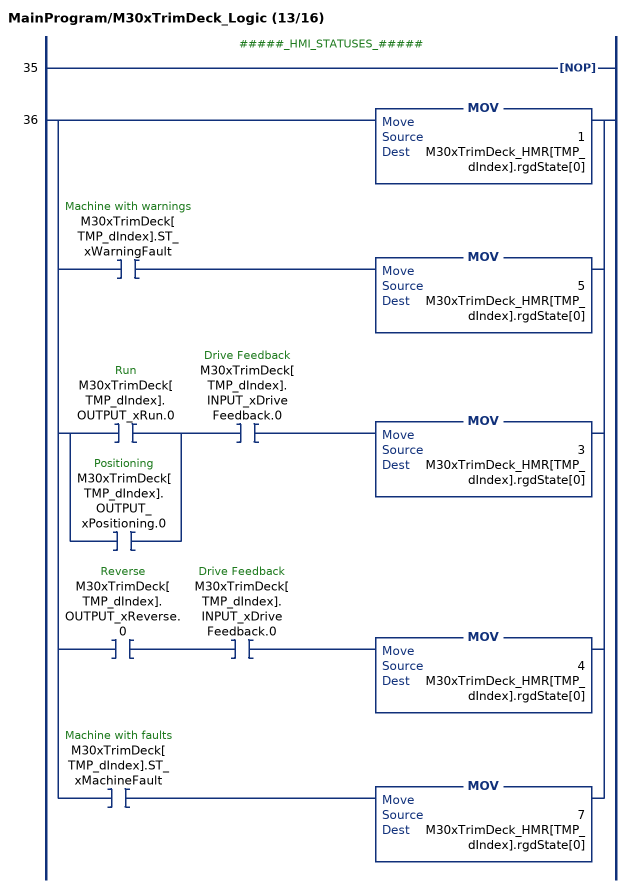
   // #####_HMI_STATUSES_#####
   35: NOP();
   36: [MOV(1,M30xTrimDeck_HMR[TMP_dIndex].rgdState[0]) ,XIC(M30xTrimDeck[TMP_dIndex].ST_xWarningFault) MOV(5,M30xTrimDeck_HMR[TMP_dIndex].rgdState[0]) ,[XIC(M30xTrimDeck[TMP_dIndex].OUTPUT_xRun.0) ,XIC(M30xTrimDeck[TMP_dIndex].OUTPUT_xPositioning.0) ] XIC(M30xTrimDeck[TMP_dIndex].INPUT_xDriveFeedback.0) MOV(3,M30xTrimDeck_HMR[TMP_dIndex].rgdState[0]) ,XIC(M30xTrimDeck[TMP_dIndex].OUTPUT_xReverse.0) XIC(M30xTrimDeck[TMP_dIndex].INPUT_xDriveFeedback.0) MOV(4,M30xTrimDeck_HMR[TMP_dIndex].rgdState[0]) ,XIC(M30xTrimDeck[TMP_dIndex].ST_xMachineFault) MOV(7,M30xTrimDeck_HMR[TMP_dIndex].rgdState[0]) ];
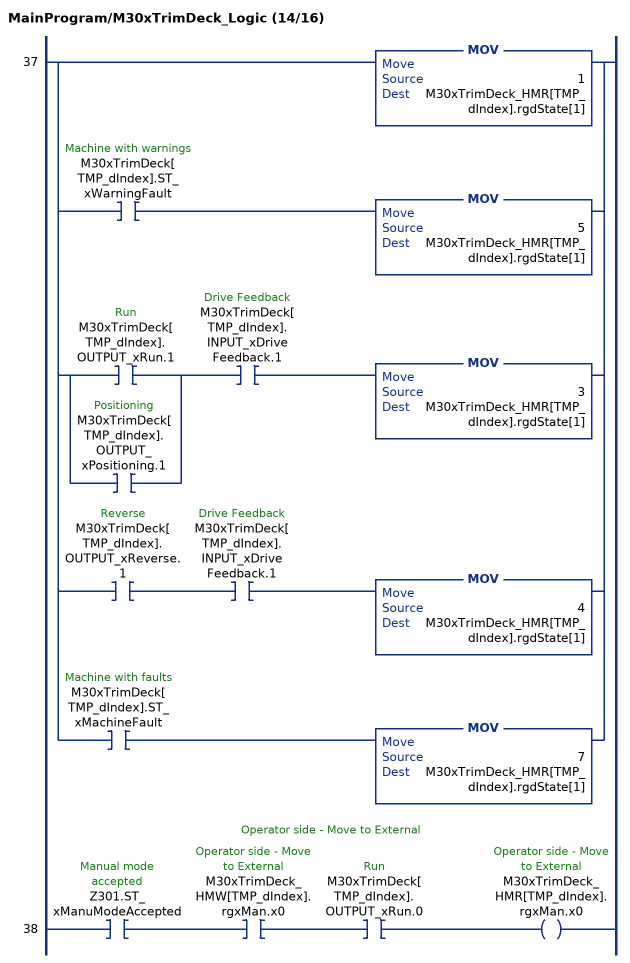
   37: [MOV(1,M30xTrimDeck_HMR[TMP_dIndex].rgdState[1]) ,XIC(M30xTrimDeck[TMP_dIndex].ST_xWarningFault) MOV(5,M30xTrimDeck_HMR[TMP_dIndex].rgdState[1]) ,[XIC(M30xTrimDeck[TMP_dIndex].OUTPUT_xRun.1) ,XIC(M30xTrimDeck[TMP_dIndex].OUTPUT_xPositioning.1) ] XIC(M30xTrimDeck[TMP_dIndex].INPUT_xDriveFeedback.1) MOV(3,M30xTrimDeck_HMR[TMP_dIndex].rgdState[1]) ,XIC(M30xTrimDeck[TMP_dIndex].OUTPUT_xReverse.1) XIC(M30xTrimDeck[TMP_dIndex].INPUT_xDriveFeedback.1) MOV(4,M30xTrimDeck_HMR[TMP_dIndex].rgdState[1]) ,XIC(M30xTrimDeck[TMP_dIndex].ST_xMachineFault) MOV(7,M30xTrimDeck_HMR[TMP_dIndex].rgdState[1]) ];
   // Operator side - Move to External
   38: XIC(Z301.ST_xManuModeAccepted)XIC(M30xTrimDeck_HMW[TMP_dIndex].rgxMan.x0)XIC(M30xTrimDeck[TMP_dIndex].OUTPUT_xRun.0)OTE(M30xTrimDeck_HMR[TMP_dIndex].rgxMan.x0);
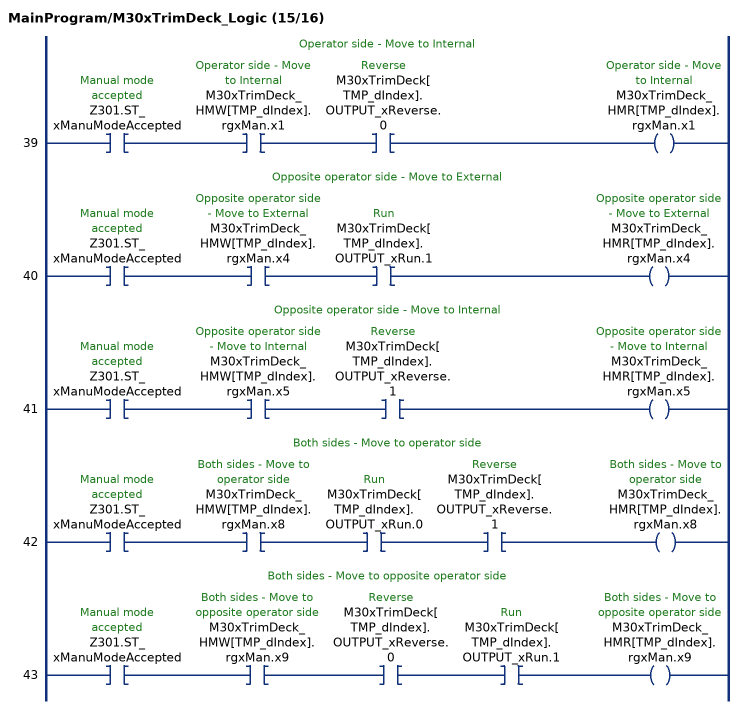
   // Operator side - Move to Internal
   39: XIC(Z301.ST_xManuModeAccepted)XIC(M30xTrimDeck_HMW[TMP_dIndex].rgxMan.x1)XIC(M30xTrimDeck[TMP_dIndex].OUTPUT_xReverse.0)OTE(M30xTrimDeck_HMR[TMP_dIndex].rgxMan.x1);
   // Opposite operator side - Move to External
   40: XIC(Z301.ST_xManuModeAccepted)XIC(M30xTrimDeck_HMW[TMP_dIndex].rgxMan.x4)XIC(M30xTrimDeck[TMP_dIndex].OUTPUT_xRun.1)OTE(M30xTrimDeck_HMR[TMP_dIndex].rgxMan.x4);
   // Opposite operator side - Move to Internal
   41: XIC(Z301.ST_xManuModeAccepted)XIC(M30xTrimDeck_HMW[TMP_dIndex].rgxMan.x5)XIC(M30xTrimDeck[TMP_dIndex].OUTPUT_xReverse.1)OTE(M30xTrimDeck_HMR[TMP_dIndex].rgxMan.x5);
   // Both sides - Move to operator side
   42: XIC(Z301.ST_xManuModeAccepted)XIC(M30xTrimDeck_HMW[TMP_dIndex].rgxMan.x8)XIC(M30xTrimDeck[TMP_dIndex].OUTPUT_xRun.0)XIC(M30xTrimDeck[TMP_dIndex].OUTPUT_xReverse.1)OTE(M30xTrimDeck_HMR[TMP_dIndex].rgxMan.x8);
   // Both sides - Move to opposite operator side
   43: XIC(Z301.ST_xManuModeAccepted)XIC(M30xTrimDeck_HMW[TMP_dIndex].rgxMan.x9)XIC(M30xTrimDeck[TMP_dIndex].OUTPUT_xReverse.0)XIC(M30xTrimDeck[TMP_dIndex].OUTPUT_xRun.1)OTE(M30xTrimDeck_HMR[TMP_dIndex].rgxMan.x9);
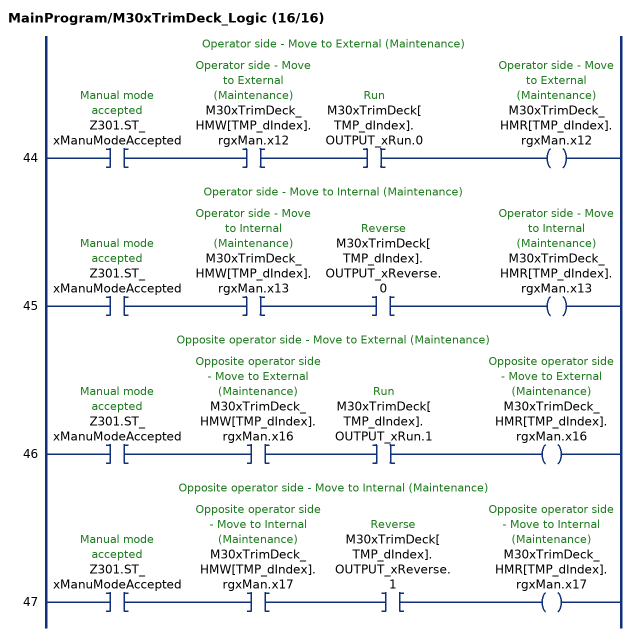
   // Operator side - Move to External (Maintenance)
   44: XIC(Z301.ST_xManuModeAccepted)XIC(M30xTrimDeck_HMW[TMP_dIndex].rgxMan.x12)XIC(M30xTrimDeck[TMP_dIndex].OUTPUT_xRun.0)OTE(M30xTrimDeck_HMR[TMP_dIndex].rgxMan.x12);
   // Operator side - Move to Internal (Maintenance)
   45: XIC(Z301.ST_xManuModeAccepted)XIC(M30xTrimDeck_HMW[TMP_dIndex].rgxMan.x13)XIC(M30xTrimDeck[TMP_dIndex].OUTPUT_xReverse.0)OTE(M30xTrimDeck_HMR[TMP_dIndex].rgxMan.x13);
   // Opposite operator side - Move to External (Maintenance)
   46: XIC(Z301.ST_xManuModeAccepted)XIC(M30xTrimDeck_HMW[TMP_dIndex].rgxMan.x16)XIC(M30xTrimDeck[TMP_dIndex].OUTPUT_xRun.1)OTE(M30xTrimDeck_HMR[TMP_dIndex].rgxMan.x16);
   // Opposite operator side - Move to Internal (Maintenance)
   47: XIC(Z301.ST_xManuModeAccepted)XIC(M30xTrimDeck_HMW[TMP_dIndex].rgxMan.x17)XIC(M30xTrimDeck[TMP_dIndex].OUTPUT_xReverse.1)OTE(M30xTrimDeck_HMR[TMP_dIndex].rgxMan.x17);
END_ROUTINE

ROUTINE M30xTrimDeckManagement   (* ladder *)
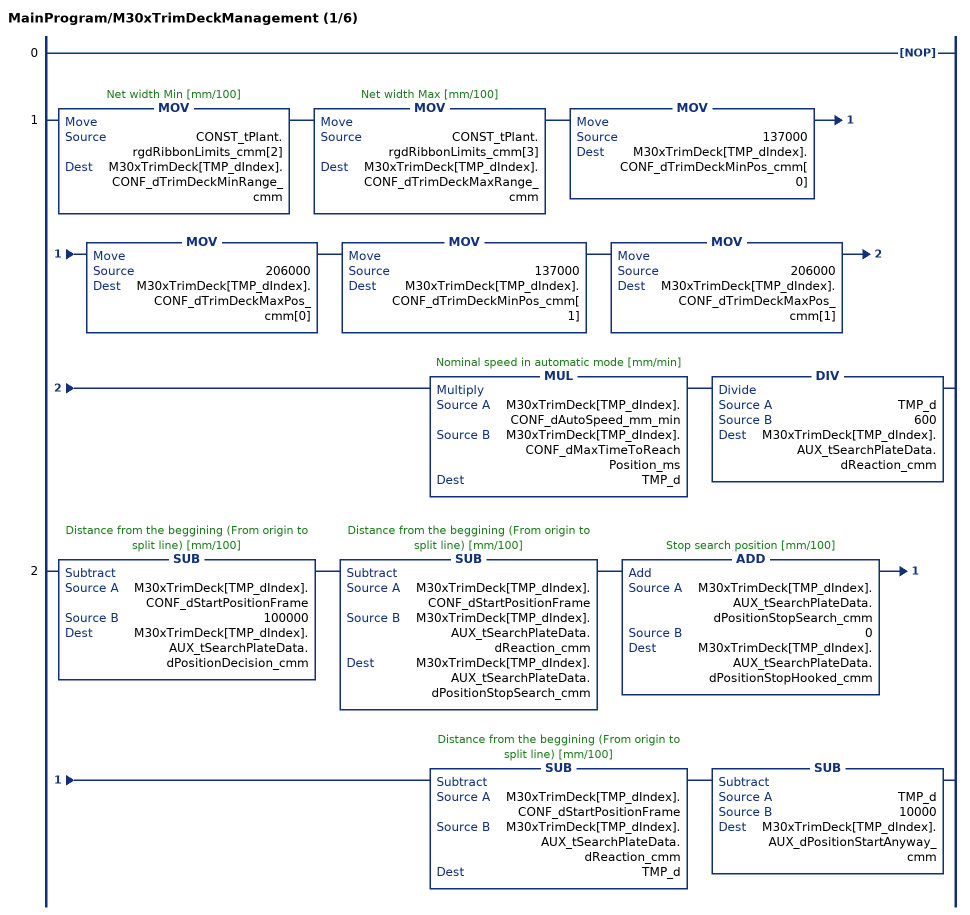
   0: NOP();
   1: MOV(CONST_tPlant.rgdRibbonLimits_cmm[2],M30xTrimDeck[TMP_dIndex].CONF_dTrimDeckMinRange_cmm)MOV(CONST_tPlant.rgdRibbonLimits_cmm[3],M30xTrimDeck[TMP_dIndex].CONF_dTrimDeckMaxRange_cmm)MOV(137000,M30xTrimDeck[TMP_dIndex].CONF_dTrimDeckMinPos_cmm[0])MOV(206000,M30xTrimDeck[TMP_dIndex].CONF_dTrimDeckMaxPos_cmm[0])MOV(137000,M30xTrimDeck[TMP_dIndex].CONF_dTrimDeckMinPos_cmm[1])MOV(206000,M30xTrimDeck[TMP_dIndex].CONF_dTrimDeckMaxPos_cmm[1])MUL(M30xTrimDeck[TMP_dIndex].CONF_dAutoSpeed_mm_min,M30xTrimDeck[TMP_dIndex].CONF_dMaxTimeToReachPosition_ms,TMP_d)DIV(TMP_d,600,M30xTrimDeck[TMP_dIndex].AUX_tSearchPlateData.dReaction_cmm);
   2: SUB(M30xTrimDeck[TMP_dIndex].CONF_dStartPositionFrame,100000,M30xTrimDeck[TMP_dIndex].AUX_tSearchPlateData.dPositionDecision_cmm)SUB(M30xTrimDeck[TMP_dIndex].CONF_dStartPositionFrame,M30xTrimDeck[TMP_dIndex].AUX_tSearchPlateData.dReaction_cmm,M30xTrimDeck[TMP_dIndex].AUX_tSearchPlateData.dPositionStopSearch_cmm)ADD(M30xTrimDeck[TMP_dIndex].AUX_tSearchPlateData.dPositionStopSearch_cmm,0,M30xTrimDeck[TMP_dIndex].AUX_tSearchPlateData.dPositionStopHooked_cmm)SUB(M30xTrimDeck[TMP_dIndex].CONF_dStartPositionFrame,M30xTrimDeck[TMP_dIndex].AUX_tSearchPlateData.dReaction_cmm,TMP_d)SUB(TMP_d,10000,M30xTrimDeck[TMP_dIndex].AUX_dPositionStartAnyway_cmm);
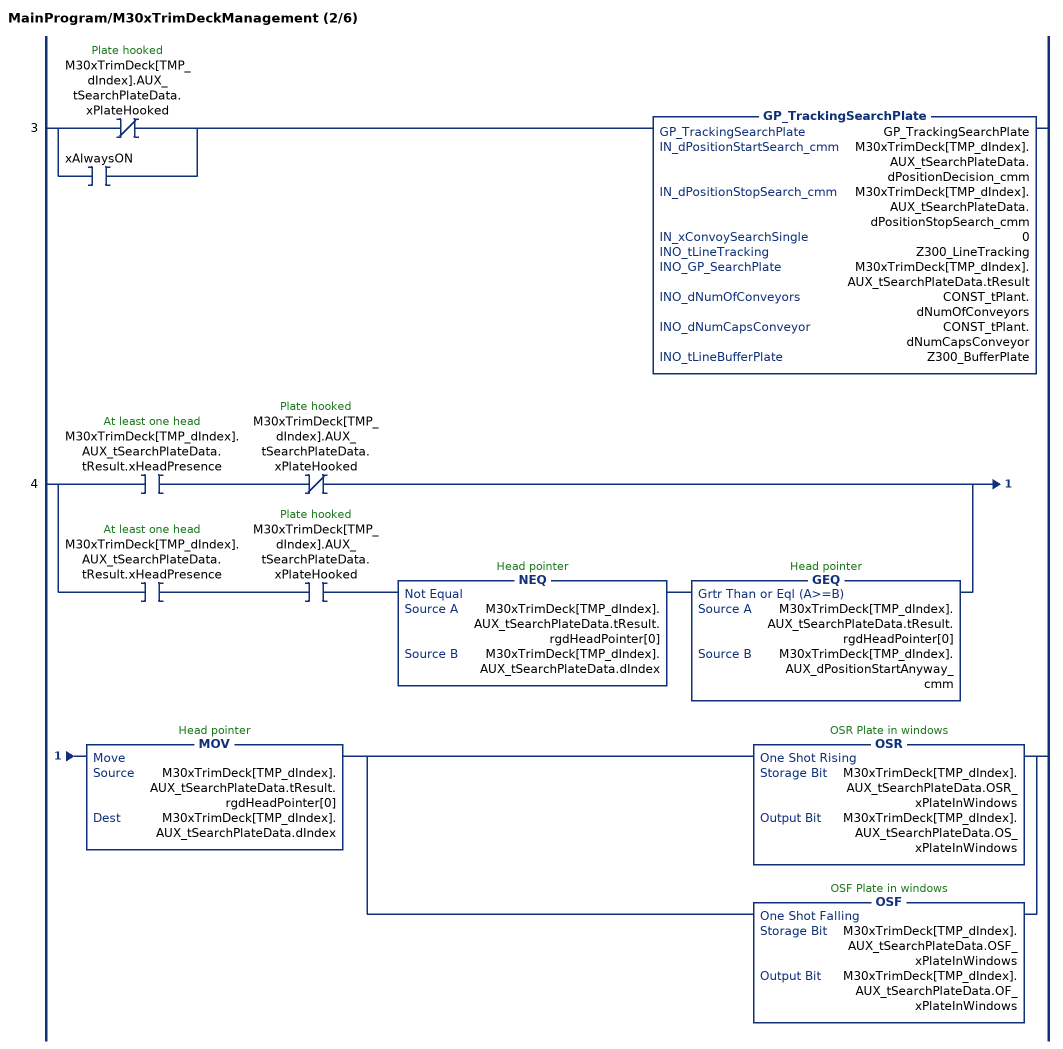
   3: [XIO(M30xTrimDeck[TMP_dIndex].AUX_tSearchPlateData.xPlateHooked) ,XIC(xAlwaysON) ]GP_TrackingSearchPlate(GP_TrackingSearchPlate,M30xTrimDeck[TMP_dIndex].AUX_tSearchPlateData.dPositionDecision_cmm,M30xTrimDeck[TMP_dIndex].AUX_tSearchPlateData.dPositionStopSearch_cmm,0,Z300_LineTracking,M30xTrimDeck[TMP_dIndex].AUX_tSearchPlateData.tResult,CONST_tPlant.dNumOfConveyors,CONST_tPlant.dNumCapsConveyor,Z300_BufferPlate);
   4: [XIC(M30xTrimDeck[TMP_dIndex].AUX_tSearchPlateData.tResult.xHeadPresence) XIO(M30xTrimDeck[TMP_dIndex].AUX_tSearchPlateData.xPlateHooked) ,XIC(M30xTrimDeck[TMP_dIndex].AUX_tSearchPlateData.tResult.xHeadPresence) XIC(M30xTrimDeck[TMP_dIndex].AUX_tSearchPlateData.xPlateHooked) NEQ(M30xTrimDeck[TMP_dIndex].AUX_tSearchPlateData.tResult.rgdHeadPointer[0],M30xTrimDeck[TMP_dIndex].AUX_tSearchPlateData.dIndex) GEQ(M30xTrimDeck[TMP_dIndex].AUX_tSearchPlateData.tResult.rgdHeadPointer[0],M30xTrimDeck[TMP_dIndex].AUX_dPositionStartAnyway_cmm) ]MOV(M30xTrimDeck[TMP_dIndex].AUX_tSearchPlateData.tResult.rgdHeadPointer[0],M30xTrimDeck[TMP_dIndex].AUX_tSearchPlateData.dIndex)[OSR(M30xTrimDeck[TMP_dIndex].AUX_tSearchPlateData.OSR_xPlateInWindows,M30xTrimDeck[TMP_dIndex].AUX_tSearchPlateData.OS_xPlateInWindows) ,OSF(M30xTrimDeck[TMP_dIndex].AUX_tSearchPlateData.OSF_xPlateInWindows,M30xTrimDeck[TMP_dIndex].AUX_tSearchPlateData.OF_xPlateInWindows) ];
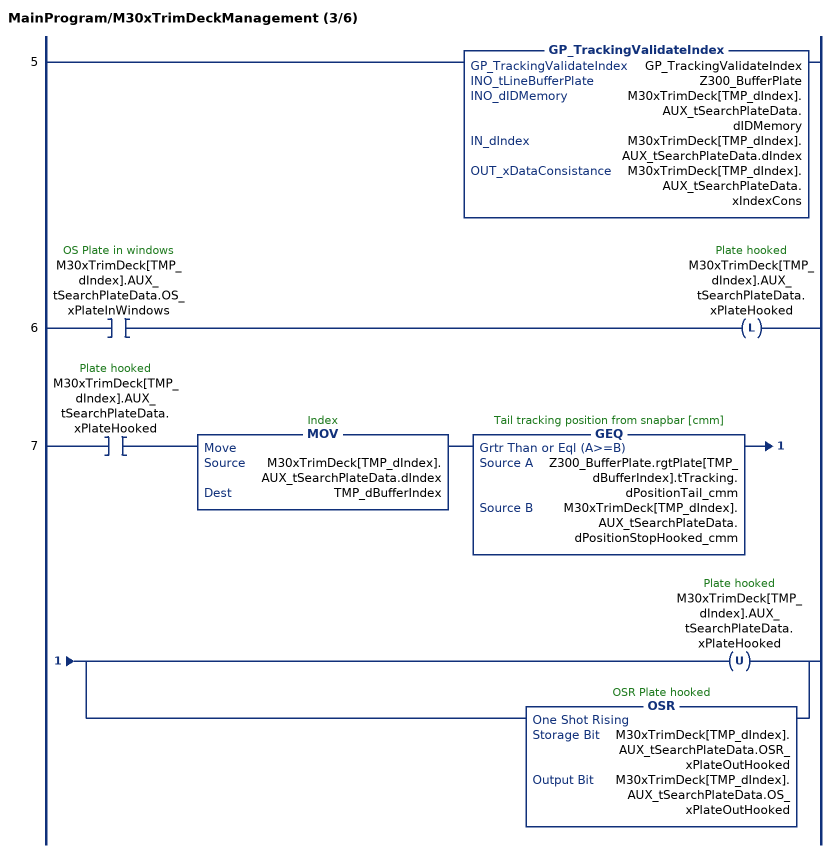
   5: GP_TrackingValidateIndex(GP_TrackingValidateIndex,Z300_BufferPlate,M30xTrimDeck[TMP_dIndex].AUX_tSearchPlateData.dIDMemory,M30xTrimDeck[TMP_dIndex].AUX_tSearchPlateData.dIndex,M30xTrimDeck[TMP_dIndex].AUX_tSearchPlateData.xIndexCons);
   6: XIC(M30xTrimDeck[TMP_dIndex].AUX_tSearchPlateData.OS_xPlateInWindows)OTL(M30xTrimDeck[TMP_dIndex].AUX_tSearchPlateData.xPlateHooked);
   7: XIC(M30xTrimDeck[TMP_dIndex].AUX_tSearchPlateData.xPlateHooked)MOV(M30xTrimDeck[TMP_dIndex].AUX_tSearchPlateData.dIndex,TMP_dBufferIndex)GEQ(Z300_BufferPlate.rgtPlate[TMP_dBufferIndex].tTracking.dPositionTail_cmm,M30xTrimDeck[TMP_dIndex].AUX_tSearchPlateData.dPositionStopHooked_cmm)[OTU(M30xTrimDeck[TMP_dIndex].AUX_tSearchPlateData.xPlateHooked) ,OSR(M30xTrimDeck[TMP_dIndex].AUX_tSearchPlateData.OSR_xPlateOutHooked,M30xTrimDeck[TMP_dIndex].AUX_tSearchPlateData.OS_xPlateOutHooked) ];
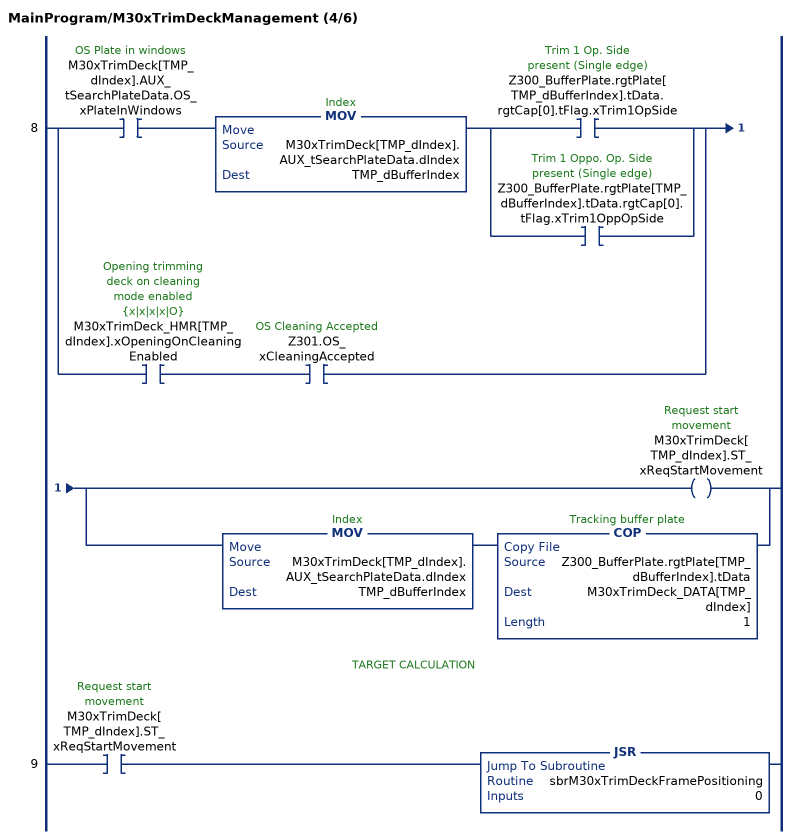
   8: [XIC(M30xTrimDeck[TMP_dIndex].AUX_tSearchPlateData.OS_xPlateInWindows) MOV(M30xTrimDeck[TMP_dIndex].AUX_tSearchPlateData.dIndex,TMP_dBufferIndex) [XIC(Z300_BufferPlate.rgtPlate[TMP_dBufferIndex].tData.rgtCap[0].tFlag.xTrim1OpSide) ,XIC(Z300_BufferPlate.rgtPlate[TMP_dBufferIndex].tData.rgtCap[0].tFlag.xTrim1OppOpSide) ] ,XIC(M30xTrimDeck_HMR[TMP_dIndex].xOpeningOnCleaningEnabled) XIC(Z301.OS_xCleaningAccepted) ][OTE(M30xTrimDeck[TMP_dIndex].ST_xReqStartMovement) ,MOV(M30xTrimDeck[TMP_dIndex].AUX_tSearchPlateData.dIndex,TMP_dBufferIndex) COP(Z300_BufferPlate.rgtPlate[TMP_dBufferIndex].tData,M30xTrimDeck_DATA[TMP_dIndex],1) ];
   // TARGET CALCULATION
   9: XIC(M30xTrimDeck[TMP_dIndex].ST_xReqStartMovement)JSR(sbrM30xTrimDeckFramePositioning,0);
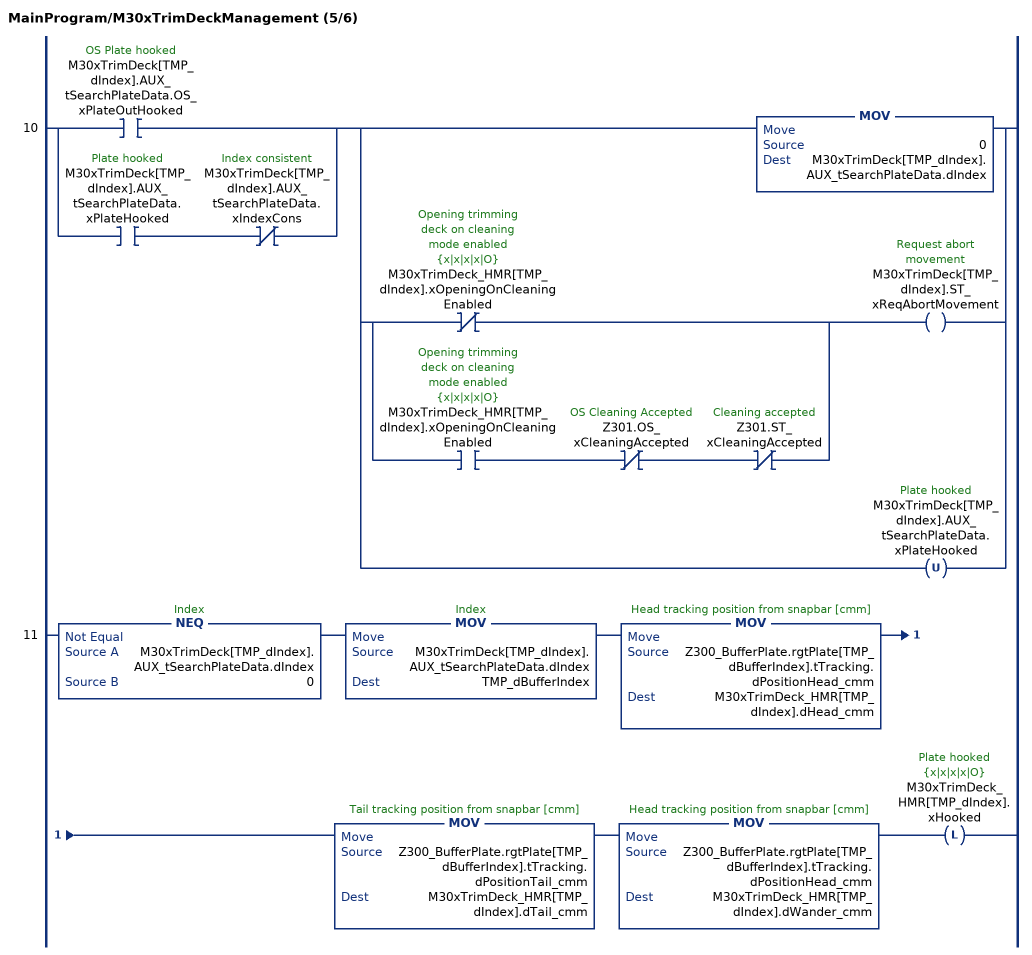
   10: [XIC(M30xTrimDeck[TMP_dIndex].AUX_tSearchPlateData.OS_xPlateOutHooked) ,XIC(M30xTrimDeck[TMP_dIndex].AUX_tSearchPlateData.xPlateHooked) XIO(M30xTrimDeck[TMP_dIndex].AUX_tSearchPlateData.xIndexCons) ][MOV(0,M30xTrimDeck[TMP_dIndex].AUX_tSearchPlateData.dIndex) ,[XIO(M30xTrimDeck_HMR[TMP_dIndex].xOpeningOnCleaningEnabled) ,XIC(M30xTrimDeck_HMR[TMP_dIndex].xOpeningOnCleaningEnabled) XIO(Z301.OS_xCleaningAccepted) XIO(Z301.ST_xCleaningAccepted) ] OTE(M30xTrimDeck[TMP_dIndex].ST_xReqAbortMovement) ,OTU(M30xTrimDeck[TMP_dIndex].AUX_tSearchPlateData.xPlateHooked) ];
   11: NEQ(M30xTrimDeck[TMP_dIndex].AUX_tSearchPlateData.dIndex,0)MOV(M30xTrimDeck[TMP_dIndex].AUX_tSearchPlateData.dIndex,TMP_dBufferIndex)MOV(Z300_BufferPlate.rgtPlate[TMP_dBufferIndex].tTracking.dPositionHead_cmm,M30xTrimDeck_HMR[TMP_dIndex].dHead_cmm)MOV(Z300_BufferPlate.rgtPlate[TMP_dBufferIndex].tTracking.dPositionTail_cmm,M30xTrimDeck_HMR[TMP_dIndex].dTail_cmm)MOV(Z300_BufferPlate.rgtPlate[TMP_dBufferIndex].tTracking.dPositionHead_cmm,M30xTrimDeck_HMR[TMP_dIndex].dWander_cmm)OTL(M30xTrimDeck_HMR[TMP_dIndex].xHooked);
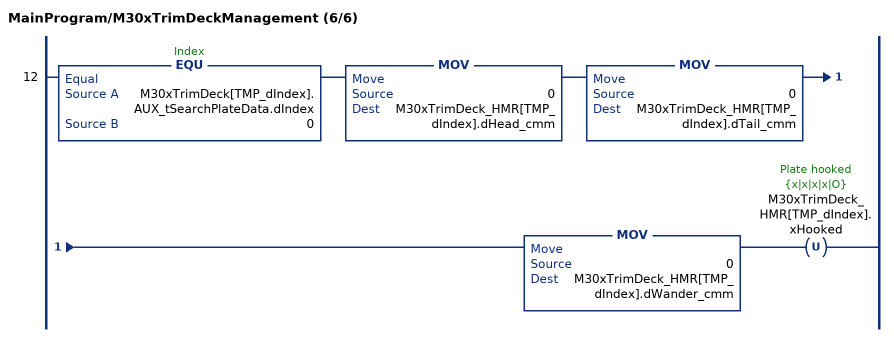
   12: EQU(M30xTrimDeck[TMP_dIndex].AUX_tSearchPlateData.dIndex,0)MOV(0,M30xTrimDeck_HMR[TMP_dIndex].dHead_cmm)MOV(0,M30xTrimDeck_HMR[TMP_dIndex].dTail_cmm)MOV(0,M30xTrimDeck_HMR[TMP_dIndex].dWander_cmm)OTU(M30xTrimDeck_HMR[TMP_dIndex].xHooked);
END_ROUTINE
